// TIA Portal project "EbAndon v2_0_1" (V15) (continued)
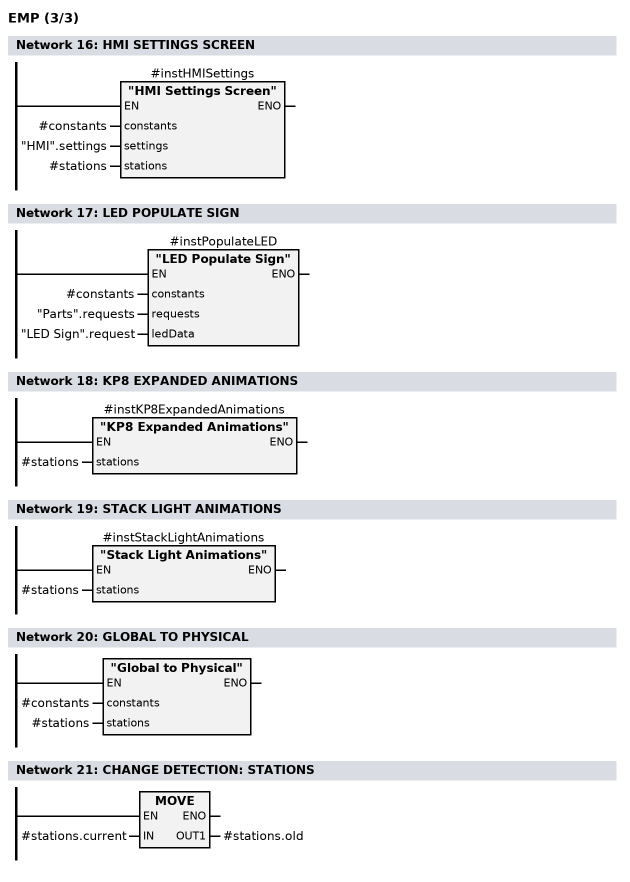
   RUNG wire#powerrail
      #instHMISettings(constants := #constants, settings := "HMI".settings, stations := #stations)
   END_RUNG
   // the same network as SCL:
   #instHMISettings(constants := #constants, settings := "HMI".settings, stations := #stations);   // "HMI Settings Screen"
END_REGION

REGION Network 17: LED POPULATE SIGN
   RUNG wire#powerrail
      #instPopulateLED(constants := #constants, requests := "Parts".requests, ledData := "LED Sign".request)
   END_RUNG
   // the same network as SCL:
   #instPopulateLED(constants := #constants, requests := "Parts".requests, ledData := "LED Sign".request);   // "LED Populate Sign"
END_REGION

REGION Network 18: KP8 EXPANDED ANIMATIONS
   RUNG wire#powerrail
      #instKP8ExpandedAnimations(stations := #stations)
   END_RUNG
   // the same network as SCL:
   #instKP8ExpandedAnimations(stations := #stations);   // "KP8 Expanded Animations"
END_REGION

REGION Network 19: STACK LIGHT ANIMATIONS
   RUNG wire#powerrail
      #instStackLightAnimations(stations := #stations)
   END_RUNG
   // the same network as SCL:
   #instStackLightAnimations(stations := #stations);   // "Stack Light Animations"
END_REGION

REGION Network 20: GLOBAL TO PHYSICAL
   RUNG wire#powerrail
      "Global to Physical"(constants := #constants, stations := #stations)
   END_RUNG
   // the same network as SCL:
   "Global to Physical"(constants := #constants, stations := #stations);
END_REGION

REGION Network 21: CHANGE DETECTION: STATIONS
   RUNG wire#powerrail
      Move(in := #stations.current, out1 => #stations.old)
   END_RUNG
   // the same network as SCL:
   #stations.old := #stations.current;
END_REGION
END_FUNCTION_BLOCK

FUNCTION_BLOCK "Code 128"   // FB2, SCL
{ S7_Optimized_Access := 'TRUE' }
VERSION : 0.1
   VAR_INPUT
      partNumber : String;
   END_VAR
   VAR_OUTPUT
      barcode : String;
   END_VAR
   VAR
      charsIn : Array[0..255] of Byte;
      charsOut : Array[0..255] of Byte;
      cnt : UInt;
      intVals : Array[0..255] of Int;
      sum : Int;
      checkSum : Int;
   END_VAR
   VAR_TEMP
      pn : String;
      i : Int;
   END_VAR
   VAR CONSTANT
      startChar : Char := 'Ì';
      stopChar : Char := 'Î';
   END_VAR
   // intVals[0] := 104;
BEGIN
   #pn := #partNumber;

   FOR #i := 0 TO 255 DO
       #charsIn[#i] := 16#00;
       #charsOut[#i] := 16#00;
       #intVals[#i] := 0;
   END_FOR;

   Strg_TO_Chars(Strg:=#pn,
                 pChars:=0,
                 Cnt=>#cnt,
                 Chars:=#charsIn);


   #sum := 104;
   FOR #i := 0 TO UINT_TO_INT(#cnt - 1) DO
       #intVals[#i] := CHAR_TO_INT(#charsIn[#i]) - 32;
       #intVals[#i] := #intVals[#i] * (#i + 1);
       #sum := #sum + #intVals[#i];
   END_FOR;
   #checkSum := (#sum MOD 103) + 32;
   IF #checkSum >= 127 THEN
       #checkSum := #checkSum + 68;
   END_IF;

   #charsOut[0] := #startChar;
   FOR #i := 1 TO UINT_TO_INT(#cnt) DO
       #charsOut[#i] := #charsIn[#i - 1];
   END_FOR;
   #charsOut[#cnt + 1] := INT_TO_BYTE(#checkSum);
   #charsOut[#cnt + 2] := INT_TO_BYTE(#stopChar);

   Chars_TO_Strg(Chars := #charsOut,
                 pChars := 0,
                 Cnt := #cnt + 3,
                 Strg => #barcode);
END_FUNCTION_BLOCK

FUNCTION_BLOCK "HMI Barcod Screen"   // FB3, SCL
{ S7_Optimized_Access := 'TRUE' }
VERSION : 0.1
   VAR_INPUT
      constants : "Constants";
   END_VAR
   VAR_IN_OUT
      partCall : "Part Call Screen";
      barcodeScreen : "Barcode Screen";
      stations : "Stations";
   END_VAR
   VAR
      address : UInt;
      button : UInt;
      instCode128 : "Code 128";
      codeOut : String;
      pnOut : WString[40];
      station : UInt;
      oldSelectedRow : Int;
      oldOrderedBtn : Bool;
   END_VAR
   VAR_TEMP
      orderCancelled : Int;
      processedPN : String[40];
      selectedPN : String[40];
      userOrdered : Bool;
      selectedRow : Int;
      position : Int;
   END_VAR
   VAR CONSTANT
      maxRows : Int := 199;
   END_VAR
BEGIN
   REGION "GET USER ROW SELECTION"
       #selectedRow := "Get Part Call Row Number"(constants := #constants,
                                                  partCall := #partCall); 
   END_REGION

   REGION "ON SELECTION OF A PART CALL ROW
       IF #selectedRow <> 0 THEN
           IF #selectedRow <> #oldSelectedRow THEN

               REGION "GET BUTTON AND STATION NUMBERS"
                   #address := #partCall.current[#selectedRow - 1].address;
                   "Address to Station and Button"(address := #address,
                                                   station => #station,
                                                   button => #button);
               END_REGION

               REGION "CONVERT STRING TO BARCODE"

                   REGION "COPY TO LOCALS"
                       #selectedPN := WSTRING_TO_STRING(#partCall.current[#selectedRow - 1].tfPartNumber.value);
                   END_REGION

                   REGION "CHECK FOR MULTI LINE"

                       REGION "GET POSITON OF CARRIAGE RETURN"
                           #position := FIND(IN1 := #selectedPN, IN2 := '$L');
                       END_REGION

                       REGION "MULTILINE"
                           IF #position <> 0 THEN
                               #processedPN := LEFT(IN := #selectedPN, L := #position - 1);
                           END_IF;
                       END_REGION

                       REGION "SINGLE LINE"
                           IF #position = 0 THEN
                               #processedPN := #selectedPN;
                           END_IF;
                       END_REGION

                   END_REGION

                   REGION "CONVERT TO BARCODE"
                       #instCode128(partNumber := #processedPN,
                                    barcode => #codeOut);
                   END_REGION

                   REGION "OUTPUT FOR HMI SCREEN"
                       #barcodeScreen.partNumber := STRING_TO_WSTRING(#processedPN);
                       #barcodeScreen.barcode := #codeOut;
                   END_REGION

               END_REGION

           END_IF;
       END_IF;
   END_REGION

   REGION "PASS USER ORDERED"

       REGION "COPY TO LOCAL"
           #userOrdered := #barcodeScreen.ordered;
       END_REGION

       REGION "TURN OFF THE LIGHTS"
           #barcodeScreen.ordered := FALSE;
       END_REGION

       REGION "ON RISING EDGE"
           IF #userOrdered AND NOT #oldOrderedBtn THEN

               REGION "SET PART ORDERED"
                   #stations.current[#station - 1].partOrdered[#button - 1] := #userOrdered;
               END_REGION

           END_IF;
       END_REGION

       REGION "CHANGE DETECTION"
           #oldOrderedBtn := #userOrdered;
       END_REGION

   END_REGION

   REGION "CHANGE DETECTION"    
       #oldSelectedRow := #selectedRow;
   END_REGION
END_FUNCTION_BLOCK

FUNCTION_BLOCK "Initialize"   // FB4, SCL
{ S7_Optimized_Access := 'TRUE' }
VERSION : 0.1
   VAR_INPUT
      constants : "Constants";
      req : Bool;
   END_VAR
   VAR_IN_OUT
      stations : "Stations";
   END_VAR
   VAR
      rtElapsed : Real;
      rt : Struct
         elapsed : LReal;
         mem : LReal;
      END_STRUCT;
   END_VAR
   VAR_TEMP
      i : Int;
      reset : Struct
         req : Bool;
         elapsed : Real;
      END_STRUCT;
      stnCount : Int;
      init : Bool;
   END_VAR
   VAR CONSTANT
      resetLimit : Real := 1.25;
   END_VAR
BEGIN
   REGION "GET STATION COUNT"
       #stnCount := #constants.stationCount - 1;
   END_REGION

   REGION "FIRST SCAN OR REQUEST"
       IF "FirstScan" OR #req THEN
           // initialize all stations on plc first scan
           FOR #i := 0 TO #stnCount DO
               #stations.current[#i].init.hard := TRUE;
           END_FOR;
       END_IF;
   END_REGION

   REGION "RUNTIME CALL"
       // get elapsed time
       #rt.elapsed := RUNTIME(#rt.mem);
       // convert to real data type
       #rtElapsed := LREAL_TO_REAL(#rt.elapsed);
   END_REGION

   REGION "BUTTON 0 BASED RESET TIMERS"
       FOR #i := 0 TO #stnCount DO

           REGION "PRE-CONDITION"
               // init off by default
               #init := FALSE;
               // request is button 0 on kp8
               #reset.req := #stations.current[#i].kp8In.%X0;
               // saved to shorter name
               #reset.elapsed := #stations.current[#i].elapsedTime.resetReq;
           END_REGION

           REGION "RESET REQUEST"
               IF NOT #reset.req THEN
                   #reset.elapsed := 0.0;
               END_IF;
               IF #reset.req THEN
                   // incriment elapsed time
                   #reset.elapsed := #reset.elapsed + #rtElapsed;
                   // timer expired condition
                   IF #reset.elapsed >= #resetLimit THEN
                       #init := TRUE;
                       #reset.elapsed := 0.0;
                   END_IF;
               END_IF;
               // save elapsed time
               #stations.current[#i].elapsedTime.resetReq := #reset.elapsed;
           END_REGION

           REGION "SAVE INITIALIZATIN REQUEST"
               #stations.current[#i].init.hard := #init;
           END_REGION

       END_FOR;
   END_REGION
END_FUNCTION_BLOCK

FUNCTION_BLOCK "Reset Init Requests"   // FB5, SCL
{ S7_Optimized_Access := 'TRUE' }
VERSION : 0.1
   VAR_INPUT
      constants : "Constants";
   END_VAR
   VAR_IN_OUT
      stations : "Stations";
   END_VAR
   VAR
      placeHolder : Bool;
   END_VAR
   VAR_TEMP
      i : Int;
      stnCount : Int;
   END_VAR
BEGIN
   REGION "GET STATION COUNT"
       #stnCount := #constants.stationCount - 1;
   END_REGION

   REGION "RESET INITIALIZATION REQUESTS
       FOR #i := 0 TO #stnCount DO
           #stations.current[#i].init.hard := FALSE;
           #stations.current[#i].init.soft := FALSE;
       END_FOR;
   END_REGION
END_FUNCTION_BLOCK

FUNCTION_BLOCK "Record Part Request"   // FB6, SCL
{ S7_Optimized_Access := 'TRUE' }
VERSION : 0.1
   VAR_INPUT
      constants : "Constants";
   END_VAR
   VAR_IN_OUT
      pRow : Int;
      requests : "Part Request Data";
      stations : "Stations";
   END_VAR
   VAR
      enterAddress : Bool;
   END_VAR
   VAR_TEMP
      address : UInt;
      hasPart : Bool;
      i : Int;
      intTime : Int;
      j : Int;
      k : Int;
      logAddress : UInt;
      noPart : Bool;
      oldPartReq : Bool;
      partReq : Bool;
      partNumber : WString;
      timeTime : Time;
      wstringTime : WString;
      stnCount : Int;
      maxReqRows : Int;
   END_VAR
BEGIN
   REGION "COPY TO LOCAL"
       #maxReqRows := #constants.partReqRows - 1;
       #stnCount := #constants.stationCount - 1;
   END_REGION

   REGION "MAIN LOOP"
       FOR #i := 0 TO #stnCount DO

           REGION "LOOP THROUGH BUTTONS"
               // j = 0 is excluded because it is used as a station reset button
               FOR #j := 1 TO 7 DO

                   REGION "PRE-CONDITION"
                       // bits for new request detection
                       #partReq := #stations.current[#i].btnStates[#j];
                       #oldPartReq := #stations.old[#i].btnStates[#j];
                   END_REGION

                   REGION "DETERMINE STATE"
                       // new request detection
                       IF #partReq AND NOT #oldPartReq THEN
                           // save to local
                           #partNumber := #stations.current[#i].partNumbers[#j];
                           // no part number
                           IF LEN(#partNumber) = 0 THEN
                               #hasPart := FALSE;
                               #noPart := TRUE;
                           END_IF;
                           // has part number
                           IF LEN(#partNumber) <> 0 THEN
                               #hasPart := TRUE;
                               #noPart := FALSE;
                           END_IF;
                       END_IF;
                   END_REGION

                   REGION "NO PART"
                       IF #noPart THEN
                           // turn off the lights
                           #hasPart := FALSE;
                           #noPart := FALSE;
                           #enterAddress := FALSE;
                       END_IF;
                   END_REGION

                   REGION "HAS PART"
                       IF #hasPart THEN
                           // turn off the lights
                           #hasPart := FALSE;
                           // calculate address
                           #address := (INT_TO_UINT(#i) + 1) * 10 + (INT_TO_UINT(#j) + 1);
                           // precondition enter address flag
                           #enterAddress := TRUE;
                           // check table for previous entry
                           FOR #k := 0 TO #maxReqRows DO
                               // save to local
                               #logAddress := #requests.row[#k].address;
                               // do not re-enter previous requests
                               IF #logAddress = #address THEN
                                   #enterAddress := FALSE;
                               END_IF;
                           END_FOR;
                       END_IF;
                   END_REGION

                   REGION "ENTER ADDRESS"
                       IF #enterAddress THEN
                           // turn off the lights
                           #enterAddress := FALSE;
                           // no processing needed
                           #requests.row[#pRow].address := #address;
                           #requests.row[#pRow].tfLine.value := #stations.current[#i].line;
                           // drop zone is unsigned so simple conversion is okay
                           #requests.row[#pRow].tfDropZone.value := USINT_TO_WSTRING(#stations.current[#i].dropZone);
                           // no processing needed
                           #requests.row[#pRow].tfPartNumber.value := #stations.current[#i].partNumbers[#j];
                           // several steps to change real to time based wstring
                           #intTime := REAL_TO_INT(#stations.current[#i].elapsedTime.partReq[#j]);
                           #timeTime := INT_TO_TIME(#intTime);
                           #wstringTime := "Time to WString"(#timeTime);
                           #requests.row[#pRow].tfTime.value := #wstringTime;
                           // incriment row pointer
                           #pRow := #pRow + 1;
                           IF #pRow > #maxReqRows THEN
                               #pRow := 0;
                           END_IF;
                       END_IF;
                   END_REGION

               END_FOR;
           END_REGION

       END_FOR;
   END_REGION
END_FUNCTION_BLOCK

FUNCTION_BLOCK "Part Timers"   // FB7, SCL
{ S7_Optimized_Access := 'TRUE' }
VERSION : 0.1
   VAR_INPUT
      constants : "Constants";
   END_VAR
   VAR_IN_OUT
      stations : "Stations";
   END_VAR
   VAR
      rt : "Runtime Data";
   END_VAR
   VAR_TEMP
      alottedTime : Real;
      btnCount : Int;
      elapsedTime : Real;
      i : Int;
      j : Int;
      partRequested : Bool;
      redTime : Real;
      remainingTime : Real;
      stnCount : Int;
      press : Struct
         current : Bool;
         old : Bool;
      END_STRUCT;
   END_VAR
BEGIN
   REGION "RUNTIME CALL"
       #rt.elapsed := RUNTIME(#rt.mem);
       #rt.asReal := LREAL_TO_REAL(#rt.elapsed);
   END_REGION

   REGION "GET STATION COUNT"
       #stnCount := #constants.stationCount - 1;
       #btnCount := #constants.buttonCount - 1;
   END_REGION

   REGION "MAIN LOOP"
       FOR #i := 0 TO #stnCount DO
           // j := 0 would be the reset button so it is skipped
           FOR #j := 1 TO #btnCount DO

               REGION "RESET PART TIMER"
                   #press.current := #stations.current[#i].btnStates[#j];
                   #press.old := #stations.old[#i].btnStates[#j];
                   IF NOT #press.current AND #press.old THEN
                           #stations.current[#i].elapsedTime.partReq[#j] := 0.0;
                   END_IF;
               END_REGION

               REGION "PART REQUEST TIMER"
                   // get and check button state 
                   #partRequested := #stations.current[#i].btnStates[#j];
                   IF #partRequested THEN

                       REGION "OUTPUT ELLAPSED TIME"
                           // get saved time
                           #elapsedTime := #stations.current[#i].elapsedTime.partReq[#j];
                           // add elapsed time
                           #elapsedTime := #elapsedTime + #rt.asReal;
                           // save new value
                           #stations.current[#i].elapsedTime.partReq[#j] := #elapsedTime;
                       END_REGION

                   END_IF;
               END_REGION

           END_FOR;
       END_FOR;
   END_REGION
END_FUNCTION_BLOCK

FUNCTION_BLOCK "Base Animations"   // FB8, SCL
{ S7_Optimized_Access := 'TRUE' }
VERSION : 0.1
   VAR_INPUT
      constants : "Constants";
   END_VAR
   VAR_IN_OUT
      stations : "Stations";
   END_VAR
   VAR_TEMP
      animation : Int;
      i : Int;
      j : Int;
      partRequested : Bool;
      partOrdered : Bool;
      elapsedTime : Real;
      criticalTime : Real;
      alottedTime : Real;
      remainingTime : Real;
      stnCount : Int;
   END_VAR
   VAR CONSTANT
      anDefault : USInt := 0;
      anRequested : USInt := 1;
      anSolidRed : USInt := 2;
      anFlashRed : USInt := 3;
      anPartOrdered : USInt := 4;
   END_VAR
BEGIN
   REGION "COPY TO LOCAL"
       #stnCount := #constants.stationCount - 1;
   END_REGION

   REGION "MAIN LOOP"
       FOR #i := 0 TO #stnCount DO
           // j := 0 would be the reset button so it is skipped
           FOR #j := 1 TO 7 DO

               REGION "PART REQUEST TIMER"

                   REGION "COPY TO LOCAL"
                       #partRequested := #stations.current[#i].btnStates[#j];
                       #partOrdered := #stations.current[#i].partOrdered[#j];
                   END_REGION

                   REGION "PART REQUESTED"
                       IF #partRequested THEN

                           REGION "COPY TO LOCAL"
                               // remaining time
                               #elapsedTime := #stations.current[#i].elapsedTime.partReq[#j];
                               #alottedTime := #stations.current[#i].presetTime.allotted[#j];
                               #remainingTime := #alottedTime - #elapsedTime;
                               // critical time
                               #criticalTime := #stations.current[#i].presetTime.critical[#j];
                           END_REGION

                           REGION "DEFAULT ANIMATION STATE"
                               IF #remainingTime > #criticalTime THEN
                                   #animation := #anRequested;
                               END_IF;
                           END_REGION

                           REGION "SOLID RED ANIMATION STATE"
                               IF #remainingTime <= #criticalTime AND #elapsedTime > 0.0 THEN
                                   #animation := #anSolidRed;
                               END_IF;
                           END_REGION

                           REGION "FLASHING RED ANIMATION STATE
                               IF #remainingTime <= 0.0 THEN
                                   #animation := #anFlashRed;
                               END_IF;
                           END_REGION ;

                           REGION "ORDERED"
                               IF #partOrdered THEN
                                   #animation := #anPartOrdered;
                               END_IF;
                           END_REGION

                       END_IF;
                   END_REGION

                   REGION "PART NOT REQUESTED"
                       IF NOT #partRequested THEN
                           #animation := #anDefault;
                       END_IF;
                   END_REGION

                   REGION "OUTPUT"
                       #stations.current[#i].animations[#j] := #animation;
                   END_REGION

               END_REGION

           END_FOR;
       END_FOR;
   END_REGION
END_FUNCTION_BLOCK

FUNCTION_BLOCK "Format Part Call Requests"   // FB9, SCL
{ S7_Optimized_Access := 'TRUE' }
VERSION : 0.1
   VAR_INPUT
      constants : "Constants";
   END_VAR
   VAR_IN_OUT
      requests : "Part Request Data";
      stations : "Stations";
   END_VAR
   VAR
      station : Int;
      button : Int;
   END_VAR
   VAR_TEMP
      address : Int;
      animate : USInt;
      maxRows : Int;
      timeAsReal : Real;
      timeAsTime : WString;
      i : Int;
      inStrRslt : Int;
      invisible : USInt;
      genericVisible : USInt;
      gray : USInt;
      darkGray : USInt;
      red : USInt;
      blue : USInt;
      redFlashing : USInt;
   END_VAR
   VAR CONSTANT
      visible : USInt := 1;
      anDefault : USInt := 0;
      anRequested : USInt := 1;
      anSolidRed : USInt := 2;
      anFlashRed : USInt := 3;
      anPartOrdered : USInt := 4;
   END_VAR
BEGIN
   REGION "COPY TO LOCAL"
       #invisible := #constants.colorLib.invisible;
       #maxRows := #constants.partReqRows - 1;
       #gray := #constants.colorLib.BgGray;
       #darkGray := #constants.colorLib.disabled;
       #blue := #constants.colorLib.BgLBl;
       #red := #constants.colorLib.BgDRd;
       #redFlashing := #constants.colorLib.FlDrd;
   END_REGION


   REGION "ITERATE THROUGH VISIBLE TABLE ROWS"
       FOR #i := 0 TO #maxRows DO

           REGION "COPY TO LOCAL"
               #address := UINT_TO_INT(#requests.row[#i].address);
           END_REGION

           REGION "HIDE UNPOPULATED ROWS"
               IF #address = 0 THEN
                   #requests.row[#i].pbSelection.animate := #invisible;
                   #requests.row[#i].rtBackground.animate := #invisible;
                   #animate := 0;
                   #requests.row[#i].tfDropZone.animate := #invisible;
                   #requests.row[#i].tfLine.animate := #invisible;
                   #requests.row[#i].tfPartNumber.animateSL := #invisible;
                   #requests.row[#i].tfPartNumber.animateDL := #invisible;
                   #requests.row[#i].tfTime.animate := #invisible;
               END_IF;
           END_REGION

           REGION "ANIMATE POPULATED ROWS"

               REGION "ANIMATE ROWS WITH DATA"
                   IF #address <> 0 THEN

                       REGION "GET POINTERS FOR STATION ARRAY"
                           #station := #address / 10 - 1;
                           #button := #address MOD 10 - 1;
                       END_REGION

                       REGION "SET ANIMATE"
                           CASE #stations.current[#station].animations[#button] OF
                               #anRequested:
                                   #animate := #gray;
                               #anSolidRed:
                                   #animate := #red;
                               #anFlashRed:
                                   #animate := #redFlashing;
                               #anPartOrdered:
                                   #animate := #blue;
                               ELSE
                                   #animate := #invisible;
                           END_CASE;
                       END_REGION


                       REGION "ANIMATIONS"

                           REGION "PUSHBUTTON VISIBILITY"
                               #requests.row[#i].pbSelection.animate := #visible;
                           END_REGION

                           REGION "BACKGROUND VISIBILITY"
                               #requests.row[#i].rtBackground.animate := #darkGray;
                           END_REGION

                           REGION "DROP ZONE" 
                               #requests.row[#i].tfDropZone.animate := #animate;
                               #requests.row[#i].tfDropZone.value := "Strip Sign"(UINT_TO_WSTRING(#stations.current[#station].dropZone));
                           END_REGION

                           REGION "LINE"
                               #requests.row[#i].tfLine.animate := #animate;
                               #requests.row[#i].tfLine.value := #stations.current[#station].line;
                           END_REGION

                           REGION "PART NUMBER"
                               #requests.row[#i].tfPartNumber.animateSL := #animate;
                               #requests.row[#i].tfPartNumber.value := #stations.current[#station].partNumbers[#button];
                               REGION "DETERMINE VISIBLE ROWS"

                                   REGION "FIND CARRIAGE RETURN"
                                       #inStrRslt := FIND(IN1 := #requests.row[#i].tfPartNumber.value,
                                                          IN2 := wstring#'$L');
                                   END_REGION

                                   REGION "SINGLE LINE"
                                       IF #inStrRslt = 0 THEN
                                           #requests.row[#i].tfPartNumber.animateSL := #animate;
                                           #requests.row[#i].tfPartNumber.animateDL := #invisible;
                                       END_IF;
                                   END_REGION

                                   REGION "DOUBLE LINE"
                                       IF #inStrRslt <> 0 THEN
                                           #requests.row[#i].tfPartNumber.animateSL := #invisible;
                                           #requests.row[#i].tfPartNumber.animateDL := #animate;
                                       END_IF;
                                   END_REGION

                               END_REGION

                           END_REGION

                           REGION "TIME"
                               #requests.row[#i].tfTime.animate := #animate;
                               #timeAsReal := #stations.current[#station].presetTime.allotted[#button];
                               #timeAsReal -= #stations.current[#station].elapsedTime.partReq[#button];
                               #requests.row[#i].tfTime.value := "Real to WString Timer"(#timeAsReal);
                           END_REGION

                       END_REGION

                   END_IF;
               END_REGION

           END_REGION

       END_FOR;
   END_REGION
END_FUNCTION_BLOCK

FUNCTION_BLOCK "KP8 Expanded Animations"   // FB10, SCL
{ S7_Optimized_Access := 'TRUE' }
VERSION : 0.1
   VAR_IN_OUT
      stations : "Stations";
   END_VAR
   VAR_TEMP
      i : Int;
      j : Int;
      colorBox : DWord;
      animation : Int;
      mask : DWord;
   END_VAR
   VAR CONSTANT
      stationCount : Int := 23;
      buttonCount : Int := 7;
      anSolidRed : USInt := 2;
      anFlashRed : USInt := 3;
      anBlue : USInt := 4;
   END_VAR
BEGIN
   REGION "LOOP THROUGH STATIONS"
       FOR #i := 0 TO #stationCount DO

           REGION "LOOP THROUGH BUTTONS"
               FOR #j := 0 TO #buttonCount DO

                   REGION "GET ANIMATION"
                       #animation := #stations.current[#i].animations[#j];
                   END_REGION

                   REGION "SOLID RED"
                       IF #animation = #anSolidRed THEN
                           #colorBox := #stations.current[#i].kp8Out;
                           #mask := 16#FEFEFEFF;
                           #mask := ROL_DWORD(IN := #mask,
                                                 N := INT_TO_UINT(#j));
                           #colorBox := #colorBox AND #mask;
                           #mask := 16#100_0000;
                           #mask := ROL_DWORD(IN := #mask,
                                                 N := INT_TO_UINT(#j));
                           #colorBox := #colorBox OR #mask;
                           #stations.current[#i].kp8Out := #colorBox;
                       END_IF;
                   END_REGION

                   REGION "FLASHING RED"
                       IF #animation = #anFlashRed THEN

                           REGION "RED ON"
                               IF "Clock_1Hz" THEN
                                   #colorBox := #stations.current[#i].kp8Out;
                                   #mask := 16#FEFEFEFF;
                                   #mask := ROL_DWORD(IN := #mask,
                                                         N := INT_TO_UINT(#j));
                                   #colorBox := #colorBox AND #mask;
                                   #mask := 16#100_0000;
                                   #mask := ROL_DWORD(IN := #mask,
                                                         N := INT_TO_UINT(#j));
                                   #colorBox := #colorBox OR #mask;
                                   #stations.current[#i].kp8Out := #colorBox;
                               END_IF;
                           END_REGION

                           REGION "RED OFF"
                               IF NOT "Clock_1Hz" THEN
                                   #colorBox := #stations.current[#i].kp8Out;
                                   #mask := 16#FEFEFEFF;
                                   #mask := ROL_DWORD(IN := #mask,
                                                         N := INT_TO_UINT(#j));
                                   #colorBox := #colorBox AND #mask;
                                   #stations.current[#i].kp8Out := #colorBox;
                               END_IF;
                           END_REGION

                       END_IF;
                   END_REGION

                   REGION "BLUE"
                       IF #animation = #anBlue THEN
                           #colorBox := #stations.current[#i].kp8Out;
                           #mask := 16#FEFEFEFF;
                           #mask := ROL_DWORD(IN := #mask,
                                              N := INT_TO_UINT(#j));
                           #colorBox := #colorBox AND #mask;
                           #mask := 16#0000_0100;
                           #mask := ROL_DWORD(IN := #mask,
                                                 N := INT_TO_UINT(#j));
                           #colorBox := #colorBox OR #mask;
                           #stations.current[#i].kp8Out := #colorBox;
                       END_IF;
                   END_REGION

               END_FOR;
           END_REGION

       END_FOR;
   END_REGION
END_FUNCTION_BLOCK

FUNCTION_BLOCK "Stack Light Animations"   // FB11, SCL
{ S7_Optimized_Access := 'TRUE' }
VERSION : 0.1
   VAR_IN_OUT
      stations : "Stations";
   END_VAR
   VAR_TEMP
      animation : Int;
      i : Int;
      j : Int;
      stackLight : DWord;
   END_VAR
   VAR CONSTANT
      anDefault : USInt := 0;
      anRequested : USInt := 1;
      anSolidRed : USInt := 2;
      anFlashRed : USInt := 3;
      anPartOrdered : USInt := 4;
      buttonCount : Int := 7;
      "Part 01" : Int := 7;
      "Part 01 Green On" : DWord := 16#0400_0000;
      "Part 01 Red On" : DWord := 16#0100_0000;
      "Part 01 Yellow On" : DWord := 16#0200_0000;
      "Part 02" : Int := 3;
      "Part 02 Green On" : DWord := 16#2000_0000;
      "Part 02 Red On" : DWord := 16#0800_0000;
      "Part 02 Yellow On" : DWord := 16#1000_0000;
      "Part 03" : Int := 6;
      "Part 03 Green On" : DWord := 16#0001_0000;
      "Part 03 Red On" : DWord := 16#4000_0000;
      "Part 03 Yellow On" : DWord := 16#8000_0000;
      "Part 04" : Int := 2;
      "Part 04 Green On" : DWord := 16#0008_0000;
      "Part 04 Yellow On" : DWord := 16#0004_0000;
      "Part 04 Red On" : DWord := 16#0002_0000;
      "Part 05" : Int := 5;
      "Part 05 Green On" : DWord := 16#0040_0000;
      "Part 05 Red On" : DWord := 16#0010_0000;
      "Part 05 Yellow On" : DWord := 16#0020_0000;
      "Part 06" : Int := 1;
      "Part 06 Green On" : DWord := 16#0000_0200;
      "Part 06 Red On" : DWord := 16#0080_0000;
      "Part 06 Yellow On" : DWord := 16#0000_0100;
      stationCount : Int := 23;
   END_VAR
BEGIN
   REGION "LOOP THROUGH STATIONS"
       FOR #i := 0 TO #stationCount DO

           REGION "LOOP THROUGH BUTTONS"
               FOR #j := 0 TO #buttonCount DO

                   REGION "COPY INTO LOCAL"
                       #stackLight := #stations.current[#i].stackLightOut;
                       #animation := #stations.current[#i].animations[#j];
                   END_REGION

                   REGION "GREEN"
                       IF #animation = #anDefault THEN
                           CASE #j OF
                               #"Part 01":
                                   #stackLight := #stackLight AND (NOT #"Part 01 Red On");
                                   #stackLight := #stackLight AND (NOT #"Part 01 Yellow On");
                                   #stackLight := #stackLight OR #"Part 01 Green On";
                               #"Part 02":
                                   #stackLight := #stackLight AND (NOT #"Part 02 Red On");
                                   #stackLight := #stackLight AND (NOT #"Part 02 Yellow On");
                                   #stackLight := #stackLight OR #"Part 02 Green On";
                               #"Part 03":
                                   #stackLight := #stackLight AND (NOT #"Part 03 Red On");
                                   #stackLight := #stackLight AND (NOT #"Part 03 Yellow On");
                                   #stackLight := #stackLight OR #"Part 03 Green On";
                               #"Part 04":
                                   #stackLight := #stackLight AND (NOT #"Part 04 Red On");
                                   #stackLight := #stackLight AND (NOT #"Part 04 Yellow On");
                                   #stackLight := #stackLight OR #"Part 04 Green On";
                               #"Part 05":
                                   #stackLight := #stackLight AND (NOT #"Part 05 Red On");
                                   #stackLight := #stackLight AND (NOT #"Part 05 Yellow On");
                                   #stackLight := #stackLight OR #"Part 05 Green On";
                               #"Part 06":
                                   #stackLight := #stackLight AND (NOT #"Part 06 Red On");
                                   #stackLight := #stackLight AND (NOT #"Part 06 Yellow On");
                                   #stackLight := #stackLight OR #"Part 06 Green On";
                               ELSE
                                   ;
                           END_CASE;
                       END_IF;
                   END_REGION

